
screen "01 Part Select" 480x800, template "Current Menu Selection"
   Button "B7" at 6,164 size 233x154; TextOff 'Text'
      on Press: function_b14e0dd5("pbs", 7)
      Visibility <- "[7]"
   Button "B6" at 6,323 size 233x154; TextOff 'Text'
      on Press: function_b14e0dd5("pbs", 6)
      Visibility <- "[6]"
   Button "B5" at 6,482 size 233x154; TextOff 'Text'
      on Press: function_b14e0dd5("pbs", 5)
      Visibility <- "[5]"
   Button "B4" at 6,641 size 233x154; TextOff 'Text'
      on Press: function_b14e0dd5("pbs", 4)
      Visibility <- "[4]"
   Button "B3" at 244,164 size 232x154; TextOff 'Text'
      on Press: function_b14e0dd5("pbs", 3)
      Visibility <- "[3]"
   Button "B2" at 244,323 size 232x154; TextOff 'Text'
      on Press: function_b14e0dd5("pbs", 2)
      Visibility <- "[2]"
   Button "B1" at 244,482 size 232x154; TextOff 'Text'
      on Press: function_b14e0dd5("pbs", 1)
      Visibility <- "[1]"
   Button "B0" at 244,641 size 232x154; TextOff 'Text'
      on Press: function_b14e0dd5("pbs", 0)
   IOField "B7 Label" at 6,164 size 233x154; FormatPattern ????????????????????????????????????????
      Appearance <- "[7]"
      ProcessValue <- "[7]"
      Visibility <- "[7]"
   IOField "B6 Label" at 6,323 size 233x154; FormatPattern ????????????????????????????????????????
      Appearance <- "[6]"
      ProcessValue <- "[6]"
      Visibility <- "[6]"
   IOField "B5 Label" at 6,482 size 233x154; FormatPattern ????????????????????????????????????????
      Appearance <- "[5]"
      ProcessValue <- "[5]"
      Visibility <- "[5]"
   IOField "B4 Label" at 6,641 size 233x154; FormatPattern ????????????????????????????????????????
      Appearance <- "[4]"
      ProcessValue <- "[4]"
      Visibility <- "[4]"
   IOField "B3 Label" at 244,164 size 232x154; FormatPattern ????????????????????????????????????????
      Appearance <- "[3]"
      ProcessValue <- "[3]"
      Visibility <- "[3]"
   IOField "B2 Label" at 244,323 size 232x154; FormatPattern ????????????????????????????????????????
      Appearance <- "[2]"
      ProcessValue <- "[2]"
      Visibility <- "[2]"
   IOField "B1 Label" at 244,482 size 232x154; FormatPattern ????????????????????????????????????????
      Appearance <- "[1]"
      ProcessValue <- "[1]"
      Visibility <- "[1]"
   IOField "B0 Label" at 244,641 size 232x154; FormatPattern ????????????????????????????????????????
      Appearance <- "[0]"
      ProcessValue <- "[0]"
      Visibility <- "[0]"

screen "02 Menu Select" 480x800, template "Current Menu Selection"
   Button "Top" at 375,164 size 100x101; TextOff 'Text'; PictureOff "basic panel top"
      on Press: function_b14e0dd5("pbs", 0)
      Appearance <- "[0]"
      Visibility <- "[0]"
   Button "Page Up" at 375,270 size 100x101; TextOff 'Text'; PictureOff "basic panel page up"
      on Press: function_b14e0dd5("pbs", 1)
      Visibility <- "[1]"
      Appearance <- "[1]"
   Button "Line Up" at 375,376 size 100x101; TextOff 'Text'; PictureOff "basic panel line up"
      on Press: function_b14e0dd5("pbs", 2)
      Appearance <- "[2]"
      Visibility <- "[2]"
   Button "Line Down" at 375,482 size 100x101; TextOff 'Text'; PictureOff "basic panel line down"
      on Press: function_b14e0dd5("pbs", 3)
      Visibility <- "[3]"
      Appearance <- "[3]"
   Button "Page Down" at 375,588 size 100x101; TextOff 'Text'; PictureOff "basic panel page down"
      on Press: function_b14e0dd5("pbs", 4)
      Appearance <- "[4]"
      Visibility <- "[4]"
   Button "Bottom" at 375,694 size 100x101; TextOff 'Text'; PictureOff "basic panel bottom"
      on Press: function_b14e0dd5("pbs", 5)
      Visibility <- "[5]"
      Appearance <- "[5]"
   IOField "brdrShortR00" at 5,164 size 365x101; FormatPattern 1
      Visibility <- "[6]"
      Appearance <- "[6]"
   IOField "brdrShortR01" at 5,270 size 365x101; FormatPattern 1
      Visibility <- "[7]"
      Appearance <- "[7]"
   IOField "brdrShortR02" at 5,376 size 365x101; FormatPattern 1
      Visibility <- "[8]"
      Appearance <- "[8]"
   IOField "brdrShortR03" at 5,482 size 365x101; FormatPattern 1
      Visibility <- "[9]"
      Appearance <- "[9]"
   IOField "brdrShortR04" at 5,588 size 365x101; FormatPattern 1
      Visibility <- "[10]"
      Appearance <- "[10]"
   IOField "brdrShortR05" at 5,694 size 365x101; FormatPattern 1
      Visibility <- "[11]"
      Appearance <- "[11]"
   Button "pbShortSelectR00" at 5,164 size 365x101; TextOff 'Text'
      on Release: ActivateScreen("01 Part Select", 0)
      on Press: function_b14e0dd5("pbs", 6)
   Button "pbShortSelectR01" at 5,270 size 365x101; TextOff 'Text'
      on Release: ActivateScreen("01 Part Select", 0)
      on Press: function_b14e0dd5("pbs", 7)
   Button "pbShortSelectR02" at 5,376 size 365x101; TextOff 'Text'
      on Release: ActivateScreen("01 Part Select", 0)
      on Press: function_b14e0dd5("pbs", 8)
   Button "pbShortSelectR03" at 5,482 size 365x101; TextOff 'Text'
      on Release: ActivateScreen("01 Part Select", 0)
      on Press: function_b14e0dd5("pbs", 9)
   Button "pbShortSelectR04" at 5,588 size 365x101; TextOff 'Text'
      on Release: ActivateScreen("01 Part Select", 0)
      on Press: function_b14e0dd5("pbs", 10)
   Button "pbShortSelectR05" at 5,694 size 365x101; TextOff 'Text'
      on Release: ActivateScreen("01 Part Select", 0)
      on Press: function_b14e0dd5("pbs", 11)
   IOField "brdrLongR00" at 5,164 size 470x101; FormatPattern 1
      Visibility <- "[18]"
   IOField "brdrLongR01" at 5,270 size 470x101; FormatPattern 1
      Visibility <- "[19]"
   IOField "brdrLongR02" at 5,376 size 470x101; FormatPattern 1
      Visibility <- "[20]"
   IOField "brdrLongR03" at 5,482 size 470x101; FormatPattern 1
      Visibility <- "[21]"
   IOField "brdrLongR04" at 5,588 size 470x101; FormatPattern 1
      Visibility <- "[22]"
   IOField "brdrLongR05" at 5,694 size 470x101; FormatPattern 1
      Visibility <- "[23]"
   Button "pbLongtSelectR00" at 5,164 size 470x101; TextOff 'Text'
      on Release: ActivateScreen("01 Part Select", 0)
      on Press: function_b14e0dd5("pbs", 6)
      Visibility <- "[18]"
   Button "pbLongtSelectR01" at 5,270 size 470x101; TextOff 'Text'
      on Release: ActivateScreen("01 Part Select", 0)
      on Press: function_b14e0dd5("pbs", 7)
      Visibility <- "[19]"
   Button "pbLongtSelectR02" at 5,376 size 470x101; TextOff 'Text'
      on Release: ActivateScreen("01 Part Select", 0)
      on Press: function_b14e0dd5("pbs", 8)
      Visibility <- "[20]"
   Button "pbLongtSelectR03" at 5,482 size 470x101; TextOff 'Text'
      on Release: ActivateScreen("01 Part Select", 0)
      on Press: function_b14e0dd5("pbs", 9)
      Visibility <- "[21]"
   Button "pbLongtSelectR04" at 5,588 size 470x101; TextOff 'Text'
      on Release: ActivateScreen("01 Part Select", 0)
      on Press: function_b14e0dd5("pbs", 10)
      Visibility <- "[22]"
   Button "pbLongtSelectR05" at 5,694 size 470x101; TextOff 'Text'
      on Release: ActivateScreen("01 Part Select", 0)
      on Press: function_b14e0dd5("pbs", 11)
      Visibility <- "[23]"
   IOField "iofLongtMenuSelectR00" at 42,166 size 430x97; FormatPattern ????????????????????????????????????????????????????????????
      Visibility <- "[18]"
      ProcessValue <- "[7]"
      Appearance <- "[18]"
   IOField "iofLongtMenuSelectR01" at 42,272 size 430x97; FormatPattern ????????????????????????????????????????????????????????????
      Visibility <- "[19]"
      ProcessValue <- "[9]"
      Appearance <- "[19]"
   IOField "iofLongtMenuSelectR02" at 42,378 size 430x97; FormatPattern ????????????????????????????????????????????????????????????
      Visibility <- "[20]"
      ProcessValue <- "[11]"
      Appearance <- "[20]"
   IOField "iofLongtMenuSelectR03" at 42,484 size 430x97; FormatPattern ????????????????????????????????????????????????????????????
      Visibility <- "[21]"
      ProcessValue <- "[13]"
      Appearance <- "[21]"
   IOField "iofLongtMenuSelectR04" at 42,590 size 430x97; FormatPattern ????????????????????????????????????????????????????????????
      Visibility <- "[22]"
      ProcessValue <- "[15]"
      Appearance <- "[22]"
   IOField "iofLongtMenuSelectR05" at 42,696 size 430x97; FormatPattern ????????????????????????????????????????????????????????????
      Visibility <- "[23]"
      ProcessValue <- "[17]"
      Appearance <- "[22]"
   IOField "iofLongLabelR00" at 7,166 size 35x97; FormatPattern ????????????????????????????????????????
      Visibility <- "[18]"
      ProcessValue <- "[6]"
      Appearance <- "[18]"
   IOField "iofLongLabelR01" at 7,272 size 35x97; FormatPattern ????????????????????????????????????????
      Appearance <- "[19]"
      ProcessValue <- "[8]"
      Visibility <- "[19]"
   IOField "iofLongLabelR02" at 7,378 size 35x97; FormatPattern ????????????????????????????????????????
      Appearance <- "[20]"
      ProcessValue <- "[10]"
      Visibility <- "[20]"
   IOField "iofLongLabelR03" at 7,484 size 35x97; FormatPattern ????????????????????????????????????????
      Appearance <- "[21]"
      ProcessValue <- "[12]"
      Visibility <- "[21]"
   IOField "iofLongLabelR04" at 7,590 size 35x97; FormatPattern ????????????????????????????????????????
      Visibility <- "[22]"
      ProcessValue <- "[14]"
      Appearance <- "[22]"
   IOField "iofLongtLabelR05" at 7,696 size 35x97; FormatPattern ????????????????????????????????????????
      Appearance <- "[23]"
      ProcessValue <- "[16]"
      Visibility <- "[23]"
   IOField "iofShortMenuSelectR00" at 42,166 size 325x97; FormatPattern ????????????????????????????????????????????????????????????
      Visibility <- "[6]"
      ProcessValue <- "[7]"
      Appearance <- "[6]"
   IOField "iofShortMenuSelectR01" at 42,272 size 325x97; FormatPattern ????????????????????????????????????????????????????????????
      Visibility <- "[7]"
      ProcessValue <- "[9]"
      Appearance <- "[7]"
   IOField "iofShortMenuSelectR02" at 42,378 size 325x97; FormatPattern ????????????????????????????????????????????????????????????
      Visibility <- "[8]"
      ProcessValue <- "[11]"
      Appearance <- "[8]"
   IOField "iofShortMenuSelectR03" at 42,484 size 325x97; FormatPattern ????????????????????????????????????????????????????????????
      Visibility <- "[9]"
      ProcessValue <- "[13]"
      Appearance <- "[9]"
   IOField "iofShortMenuSelectR04" at 42,590 size 325x97; FormatPattern ????????????????????????????????????????????????????????????
      Visibility <- "[10]"
      ProcessValue <- "[15]"
      Appearance <- "[10]"
   IOField "iofShortMenuSelectR05" at 42,696 size 325x97; FormatPattern ????????????????????????????????????????????????????????????
      Visibility <- "[11]"
      ProcessValue <- "[17]"
      Appearance <- "[11]"
   IOField "iofShortLabelR00" at 7,166 size 35x97; FormatPattern ????????????????????????????????????????
      Appearance <- "[6]"
      ProcessValue <- "[6]"
      Visibility <- "[6]"
   IOField "iofShortLabelR01" at 7,272 size 35x97; FormatPattern ????????????????????????????????????????
      Appearance <- "[7]"
      ProcessValue <- "[8]"
      Visibility <- "[7]"
   IOField "iofShortLabelR02" at 7,378 size 35x97; FormatPattern ????????????????????????????????????????
      Appearance <- "[8]"
      ProcessValue <- "[10]"
      Visibility <- "[8]"
   IOField "iofShortLabelR03" at 7,484 size 35x97; FormatPattern ????????????????????????????????????????
      Appearance <- "[9]"
      ProcessValue <- "[12]"
      Visibility <- "[9]"
   IOField "iofShortLabelR04" at 7,590 size 35x97; FormatPattern ????????????????????????????????????????
      Appearance <- "[10]"
      ProcessValue <- "[14]"
      Visibility <- "[10]"
   IOField "iofShorttLabelR05" at 7,696 size 35x97; FormatPattern ????????????????????????????????????????
      Appearance <- "[11]"
      ProcessValue <- "[16]"
      Visibility <- "[11]"

Template "Current Menu Selection" 480x800
   IOField "Menu Select Label" at 6,5 size 470x154; FormatPattern ????????????????????????????????????????????????????????????
      Appearance <- "[0]"
      Visibility <- "[0]"
      ProcessValue <- "[0]"
   Button "PB Menu Select" at 6,5 size 470x154; TextOff 'Text'
      on Release: ActivateScreen("02 Menu Select", 0)
      on Press: function_b14e0dd5("pb", 0)
*)

(* ===== HMI "HMI_RT_6" =====
system functions are stored by id; their names below are inferred from use
connection "cv01": ETHERNET, SMART_S7_1500_OMS

HMI tags "Default tag table"
   "station" : HMIS: Compressed = PLC "HMI Stations".me[0] AT %DB1.DBW0, 100 ms

screen "01 Part Select" 480x800, template "Current Menu Selection"
   Button "B7" at 6,164 size 233x154; TextOff 'Text'
      on Press: function_b14e0dd5("pbs", 7)
      Visibility <- "[7]"
   Button "B6" at 6,323 size 233x154; TextOff 'Text'
      on Press: function_b14e0dd5("pbs", 6)
      Visibility <- "[6]"
   Button "B5" at 6,482 size 233x154; TextOff 'Text'
      on Press: function_b14e0dd5("pbs", 5)
      Visibility <- "[5]"
   Button "B4" at 6,641 size 233x154; TextOff 'Text'
      on Press: function_b14e0dd5("pbs", 4)
      Visibility <- "[4]"
   Button "B3" at 244,164 size 232x154; TextOff 'Text'
      on Press: function_b14e0dd5("pbs", 3)
      Visibility <- "[3]"
   Button "B2" at 244,323 size 232x154; TextOff 'Text'
      on Press: function_b14e0dd5("pbs", 2)
      Visibility <- "[2]"
   Button "B1" at 244,482 size 232x154; TextOff 'Text'
      on Press: function_b14e0dd5("pbs", 1)
      Visibility <- "[1]"
   Button "B0" at 244,641 size 232x154; TextOff 'Text'
      on Press: function_b14e0dd5("pbs", 0)
   IOField "B7 Label" at 6,164 size 233x154; FormatPattern ????????????????????????????????????????
      Appearance <- "[7]"
      ProcessValue <- "[7]"
      Visibility <- "[7]"
   IOField "B6 Label" at 6,323 size 233x154; FormatPattern ????????????????????????????????????????
      Appearance <- "[6]"
      ProcessValue <- "[6]"
      Visibility <- "[6]"
   IOField "B5 Label" at 6,482 size 233x154; FormatPattern ????????????????????????????????????????
      Appearance <- "[5]"
      ProcessValue <- "[5]"
      Visibility <- "[5]"
   IOField "B4 Label" at 6,641 size 233x154; FormatPattern ????????????????????????????????????????
      Appearance <- "[4]"
      ProcessValue <- "[4]"
      Visibility <- "[4]"
   IOField "B3 Label" at 244,164 size 232x154; FormatPattern ????????????????????????????????????????
      Appearance <- "[3]"
      ProcessValue <- "[3]"
      Visibility <- "[3]"
   IOField "B2 Label" at 244,323 size 232x154; FormatPattern ????????????????????????????????????????
      Appearance <- "[2]"
      ProcessValue <- "[2]"
      Visibility <- "[2]"
   IOField "B1 Label" at 244,482 size 232x154; FormatPattern ????????????????????????????????????????
      Appearance <- "[1]"
      ProcessValue <- "[1]"
      Visibility <- "[1]"
   IOField "B0 Label" at 244,641 size 232x154; FormatPattern ????????????????????????????????????????
      Appearance <- "[0]"
      ProcessValue <- "[0]"
      Visibility <- "[0]"
   TextField "B7 BG" at 6,164 size 233x154; Text '1'

screen "02 Menu Select" 480x800, template "Current Menu Selection"
   Button "Top" at 375,164 size 100x101; TextOff 'Text'; PictureOff "basic panel top"
      on Press: function_b14e0dd5("pbs", 0)
      Appearance <- "[0]"
      Visibility <- "[0]"
   Button "Page Up" at 375,270 size 100x101; TextOff 'Text'; PictureOff "basic panel page up"
      on Press: function_b14e0dd5("pbs", 1)
      Visibility <- "[1]"
      Appearance <- "[1]"
   Button "Line Up" at 375,376 size 100x101; TextOff 'Text'; PictureOff "basic panel line up"
      on Press: function_b14e0dd5("pbs", 2)
      Appearance <- "[2]"
      Visibility <- "[2]"
   Button "Line Down" at 375,482 size 100x101; TextOff 'Text'; PictureOff "basic panel line down"
      on Press: function_b14e0dd5("pbs", 3)
      Visibility <- "[3]"
      Appearance <- "[3]"
   Button "Page Down" at 375,588 size 100x101; TextOff 'Text'; PictureOff "basic panel page down"
      on Press: function_b14e0dd5("pbs", 4)
      Appearance <- "[4]"
      Visibility <- "[4]"
   Button "Bottom" at 375,694 size 100x101; TextOff 'Text'; PictureOff "basic panel bottom"
      on Press: function_b14e0dd5("pbs", 5)
      Visibility <- "[5]"
      Appearance <- "[5]"
   IOField "brdrShortR00" at 5,164 size 365x101; FormatPattern 1
      Visibility <- "[6]"
      Appearance <- "[6]"
   IOField "brdrShortR01" at 5,270 size 365x101; FormatPattern 1
      Visibility <- "[7]"
      Appearance <- "[7]"
   IOField "brdrShortR02" at 5,376 size 365x101; FormatPattern 1
      Visibility <- "[8]"
      Appearance <- "[8]"
   IOField "brdrShortR03" at 5,482 size 365x101; FormatPattern 1
      Visibility <- "[9]"
      Appearance <- "[9]"
   IOField "brdrShortR04" at 5,588 size 365x101; FormatPattern 1
      Visibility <- "[10]"
      Appearance <- "[10]"
   IOField "brdrShortR05" at 5,694 size 365x101; FormatPattern 1
      Visibility <- "[11]"
      Appearance <- "[11]"
   Button "pbShortSelectR00" at 5,164 size 365x101; TextOff 'Text'
      on Release: ActivateScreen("01 Part Select", 0)
      on Press: function_b14e0dd5("pbs", 6)
   Button "pbShortSelectR01" at 5,270 size 365x101; TextOff 'Text'
      on Release: ActivateScreen("01 Part Select", 0)
      on Press: function_b14e0dd5("pbs", 7)
   Button "pbShortSelectR02" at 5,376 size 365x101; TextOff 'Text'
      on Release: ActivateScreen("01 Part Select", 0)
      on Press: function_b14e0dd5("pbs", 8)
   Button "pbShortSelectR03" at 5,482 size 365x101; TextOff 'Text'
      on Release: ActivateScreen("01 Part Select", 0)
      on Press: function_b14e0dd5("pbs", 9)
   Button "pbShortSelectR04" at 5,588 size 365x101; TextOff 'Text'
      on Release: ActivateScreen("01 Part Select", 0)
      on Press: function_b14e0dd5("pbs", 10)
   Button "pbShortSelectR05" at 5,694 size 365x101; TextOff 'Text'
      on Release: ActivateScreen("01 Part Select", 0)
      on Press: function_b14e0dd5("pbs", 11)
   IOField "brdrLongR00" at 5,164 size 470x101; FormatPattern 1
      Visibility <- "[18]"
   IOField "brdrLongR01" at 5,270 size 470x101; FormatPattern 1
      Visibility <- "[19]"
   IOField "brdrLongR02" at 5,376 size 470x101; FormatPattern 1
      Visibility <- "[20]"
   IOField "brdrLongR03" at 5,482 size 470x101; FormatPattern 1
      Visibility <- "[21]"
   IOField "brdrLongR04" at 5,588 size 470x101; FormatPattern 1
      Visibility <- "[22]"
   IOField "brdrLongR05" at 5,694 size 470x101; FormatPattern 1
      Visibility <- "[23]"
   Button "pbLongtSelectR00" at 5,164 size 470x101; TextOff 'Text'
      on Release: ActivateScreen("01 Part Select", 0)
      on Press: function_b14e0dd5("pbs", 6)
      Visibility <- "[18]"
   Button "pbLongtSelectR01" at 5,270 size 470x101; TextOff 'Text'
      on Release: ActivateScreen("01 Part Select", 0)
      on Press: function_b14e0dd5("pbs", 7)
      Visibility <- "[19]"
   Button "pbLongtSelectR02" at 5,376 size 470x101; TextOff 'Text'
      on Release: ActivateScreen("01 Part Select", 0)
      on Press: function_b14e0dd5("pbs", 8)
      Visibility <- "[20]"
   Button "pbLongtSelectR03" at 5,482 size 470x101; TextOff 'Text'
      on Release: ActivateScreen("01 Part Select", 0)
      on Press: function_b14e0dd5("pbs", 9)
      Visibility <- "[21]"
   Button "pbLongtSelectR04" at 5,588 size 470x101; TextOff 'Text'
      on Release: ActivateScreen("01 Part Select", 0)
      on Press: function_b14e0dd5("pbs", 10)
      Visibility <- "[22]"
   Button "pbLongtSelectR05" at 5,694 size 470x101; TextOff 'Text'
      on Release: ActivateScreen("01 Part Select", 0)
      on Press: function_b14e0dd5("pbs", 11)
      Visibility <- "[23]"
   IOField "iofLongtMenuSelectR00" at 42,166 size 430x97; FormatPattern ????????????????????????????????????????????????????????????
      Visibility <- "[18]"
      ProcessValue <- "[7]"
      Appearance <- "[18]"
   IOField "iofLongtMenuSelectR01" at 42,272 size 430x97; FormatPattern ????????????????????????????????????????????????????????????
      Visibility <- "[19]"
      ProcessValue <- "[9]"
      Appearance <- "[19]"
   IOField "iofLongtMenuSelectR02" at 42,378 size 430x97; FormatPattern ????????????????????????????????????????????????????????????
      Visibility <- "[20]"
      ProcessValue <- "[11]"
      Appearance <- "[20]"
   IOField "iofLongtMenuSelectR03" at 42,484 size 430x97; FormatPattern ????????????????????????????????????????????????????????????
      Visibility <- "[21]"
      ProcessValue <- "[13]"
      Appearance <- "[21]"
   IOField "iofLongtMenuSelectR04" at 42,590 size 430x97; FormatPattern ????????????????????????????????????????????????????????????
      Visibility <- "[22]"
      ProcessValue <- "[15]"
      Appearance <- "[22]"
   IOField "iofLongtMenuSelectR05" at 42,696 size 430x97; FormatPattern ????????????????????????????????????????????????????????????
      Visibility <- "[23]"
      ProcessValue <- "[17]"
      Appearance <- "[22]"
   IOField "iofLongLabelR00" at 7,166 size 35x97; FormatPattern ????????????????????????????????????????
      Visibility <- "[18]"
      ProcessValue <- "[6]"
      Appearance <- "[18]"
   IOField "iofLongLabelR01" at 7,272 size 35x97; FormatPattern ????????????????????????????????????????
      Appearance <- "[19]"
      ProcessValue <- "[8]"
      Visibility <- "[19]"
   IOField "iofLongLabelR02" at 7,378 size 35x97; FormatPattern ????????????????????????????????????????
      Appearance <- "[20]"
      ProcessValue <- "[10]"
      Visibility <- "[20]"
   IOField "iofLongLabelR03" at 7,484 size 35x97; FormatPattern ????????????????????????????????????????
      Appearance <- "[21]"
      ProcessValue <- "[12]"
      Visibility <- "[21]"
   IOField "iofLongLabelR04" at 7,590 size 35x97; FormatPattern ????????????????????????????????????????
      Visibility <- "[22]"
      ProcessValue <- "[14]"
      Appearance <- "[22]"
   IOField "iofLongtLabelR05" at 7,696 size 35x97; FormatPattern ????????????????????????????????????????
      Appearance <- "[23]"
      ProcessValue <- "[16]"
      Visibility <- "[23]"
   IOField "iofShortMenuSelectR00" at 42,166 size 325x97; FormatPattern ????????????????????????????????????????????????????????????
      Visibility <- "[6]"
      ProcessValue <- "[7]"
      Appearance <- "[6]"
   IOField "iofShortMenuSelectR01" at 42,272 size 325x97; FormatPattern ????????????????????????????????????????????????????????????
      Visibility <- "[7]"
      ProcessValue <- "[9]"
      Appearance <- "[7]"
   IOField "iofShortMenuSelectR02" at 42,378 size 325x97; FormatPattern ????????????????????????????????????????????????????????????
      Visibility <- "[8]"
      ProcessValue <- "[11]"
      Appearance <- "[8]"
   IOField "iofShortMenuSelectR03" at 42,484 size 325x97; FormatPattern ????????????????????????????????????????????????????????????
      Visibility <- "[9]"
      ProcessValue <- "[13]"
      Appearance <- "[9]"
   IOField "iofShortMenuSelectR04" at 42,590 size 325x97; FormatPattern ????????????????????????????????????????????????????????????
      Visibility <- "[10]"
      ProcessValue <- "[15]"
      Appearance <- "[10]"
   IOField "iofShortMenuSelectR05" at 42,696 size 325x97; FormatPattern ????????????????????????????????????????????????????????????
      Visibility <- "[11]"
      ProcessValue <- "[17]"
      Appearance <- "[11]"
   IOField "iofShortLabelR00" at 7,166 size 35x97; FormatPattern ????????????????????????????????????????
      Appearance <- "[6]"
      ProcessValue <- "[6]"
      Visibility <- "[6]"
   IOField "iofShortLabelR01" at 7,272 size 35x97; FormatPattern ????????????????????????????????????????
      Appearance <- "[7]"
      ProcessValue <- "[8]"
      Visibility <- "[7]"
   IOField "iofShortLabelR02" at 7,378 size 35x97; FormatPattern ????????????????????????????????????????
      Appearance <- "[8]"
      ProcessValue <- "[10]"
      Visibility <- "[8]"
   IOField "iofShortLabelR03" at 7,484 size 35x97; FormatPattern ????????????????????????????????????????
      Appearance <- "[9]"
      ProcessValue <- "[12]"
      Visibility <- "[9]"
   IOField "iofShortLabelR04" at 7,590 size 35x97; FormatPattern ????????????????????????????????????????
      Appearance <- "[10]"
      ProcessValue <- "[14]"
      Visibility <- "[10]"
   IOField "iofShorttLabelR05" at 7,696 size 35x97; FormatPattern ????????????????????????????????????????
      Appearance <- "[11]"
      ProcessValue <- "[16]"
      Visibility <- "[11]"

Template "Current Menu Selection" 480x800
   IOField "Menu Select Label" at 6,5 size 470x154; FormatPattern ????????????????????????????????????????????????????????????
      Appearance <- "[0]"
      Visibility <- "[0]"
      ProcessValue <- "[0]"
   Button "PB Menu Select" at 6,5 size 470x154; TextOff 'Text'
      on Release: ActivateScreen("02 Menu Select", 0)
      on Press: function_b14e0dd5("pb", 0)
*)

(* ===== HMI "HMI_RT_7" =====
system functions are stored by id; their names below are inferred from use
connection "pc01": ETHERNET, SMART_S7_1500_OMS

HMI tags "Default tag table"
   "station" : HMIS: Compressed = PLC "HMI Stations".me[4] AT %DB1.DBW0, 100 ms

screen "01 Part Select" 480x800, template "Current Menu Selection"
   Button "B7" at 6,164 size 233x154; TextOff 'Text'
      on Press: function_b14e0dd5("pbs", 7)
      Visibility <- "[7]"
   Button "B6" at 6,323 size 233x154; TextOff 'Text'
      on Press: function_b14e0dd5("pbs", 6)
      Visibility <- "[6]"
   Button "B5" at 6,482 size 233x154; TextOff 'Text'
      on Press: function_b14e0dd5("pbs", 5)
      Visibility <- "[5]"
   Button "B4" at 6,641 size 233x154; TextOff 'Text'
      on Press: function_b14e0dd5("pbs", 4)
      Visibility <- "[4]"
   Button "B3" at 244,164 size 232x154; TextOff 'Text'
      on Press: function_b14e0dd5("pbs", 3)
      Visibility <- "[3]"
   Button "B2" at 244,323 size 232x154; TextOff 'Text'
      on Press: function_b14e0dd5("pbs", 2)
      Visibility <- "[2]"
   Button "B1" at 244,482 size 232x154; TextOff 'Text'
      on Press: function_b14e0dd5("pbs", 1)
      Visibility <- "[1]"
   Button "B0" at 244,641 size 232x154; TextOff 'Text'
      on Press: function_b14e0dd5("pbs", 0)
   IOField "B7 Label" at 6,164 size 233x154; FormatPattern ????????????????????????????????????????
      Appearance <- "[7]"
      ProcessValue <- "[7]"
      Visibility <- "[7]"
   IOField "B6 Label" at 6,323 size 233x154; FormatPattern ????????????????????????????????????????
      Appearance <- "[6]"
      ProcessValue <- "[6]"
      Visibility <- "[6]"
   IOField "B5 Label" at 6,482 size 233x154; FormatPattern ????????????????????????????????????????
      Appearance <- "[5]"
      ProcessValue <- "[5]"
      Visibility <- "[5]"
   IOField "B4 Label" at 6,641 size 233x154; FormatPattern ????????????????????????????????????????
      Appearance <- "[4]"
      ProcessValue <- "[4]"
      Visibility <- "[4]"
   IOField "B3 Label" at 244,164 size 232x154; FormatPattern ????????????????????????????????????????
      Appearance <- "[3]"
      ProcessValue <- "[3]"
      Visibility <- "[3]"
   IOField "B2 Label" at 244,323 size 232x154; FormatPattern ????????????????????????????????????????
      Appearance <- "[2]"
      ProcessValue <- "[2]"
      Visibility <- "[2]"
   IOField "B1 Label" at 244,482 size 232x154; FormatPattern ????????????????????????????????????????
      Appearance <- "[1]"
      ProcessValue <- "[1]"
      Visibility <- "[1]"
   IOField "B0 Label" at 244,641 size 232x154; FormatPattern ????????????????????????????????????????
      Appearance <- "[0]"
      ProcessValue <- "[0]"
      Visibility <- "[0]"

screen "02 Menu Select" 480x800, template "Current Menu Selection"
   Button "Top" at 375,164 size 100x101; TextOff 'Text'; PictureOff "basic panel top"
      on Press: function_b14e0dd5("pbs", 0)
      Appearance <- "[0]"
      Visibility <- "[0]"
   Button "Page Up" at 375,270 size 100x101; TextOff 'Text'; PictureOff "basic panel page up"
      on Press: function_b14e0dd5("pbs", 1)
      Visibility <- "[1]"
      Appearance <- "[1]"
   Button "Line Up" at 375,376 size 100x101; TextOff 'Text'; PictureOff "basic panel line up"
      on Press: function_b14e0dd5("pbs", 2)
      Appearance <- "[2]"
      Visibility <- "[2]"
   Button "Line Down" at 375,482 size 100x101; TextOff 'Text'; PictureOff "basic panel line down"
      on Press: function_b14e0dd5("pbs", 3)
      Visibility <- "[3]"
      Appearance <- "[3]"
   Button "Page Down" at 375,588 size 100x101; TextOff 'Text'; PictureOff "basic panel page down"
      on Press: function_b14e0dd5("pbs", 4)
      Appearance <- "[4]"
      Visibility <- "[4]"
   Button "Bottom" at 375,694 size 100x101; TextOff 'Text'; PictureOff "basic panel bottom"
      on Press: function_b14e0dd5("pbs", 5)
      Visibility <- "[5]"
      Appearance <- "[5]"
   IOField "brdrShortR00" at 5,164 size 365x101; FormatPattern 1
      Visibility <- "[6]"
      Appearance <- "[6]"
   IOField "brdrShortR01" at 5,270 size 365x101; FormatPattern 1
      Visibility <- "[7]"
      Appearance <- "[7]"
   IOField "brdrShortR02" at 5,376 size 365x101; FormatPattern 1
      Visibility <- "[8]"
      Appearance <- "[8]"
   IOField "brdrShortR03" at 5,482 size 365x101; FormatPattern 1
      Visibility <- "[9]"
      Appearance <- "[9]"
   IOField "brdrShortR04" at 5,588 size 365x101; FormatPattern 1
      Visibility <- "[10]"
      Appearance <- "[10]"
   IOField "brdrShortR05" at 5,694 size 365x101; FormatPattern 1
      Visibility <- "[11]"
      Appearance <- "[11]"
   Button "pbShortSelectR00" at 5,164 size 365x101; TextOff 'Text'
      on Release: ActivateScreen("01 Part Select", 0)
      on Press: function_b14e0dd5("pbs", 6)
   Button "pbShortSelectR01" at 5,270 size 365x101; TextOff 'Text'
      on Release: ActivateScreen("01 Part Select", 0)
      on Press: function_b14e0dd5("pbs", 7)
   Button "pbShortSelectR02" at 5,376 size 365x101; TextOff 'Text'
      on Release: ActivateScreen("01 Part Select", 0)
      on Press: function_b14e0dd5("pbs", 8)
   Button "pbShortSelectR03" at 5,482 size 365x101; TextOff 'Text'
      on Release: ActivateScreen("01 Part Select", 0)
      on Press: function_b14e0dd5("pbs", 9)
   Button "pbShortSelectR04" at 5,588 size 365x101; TextOff 'Text'
      on Release: ActivateScreen("01 Part Select", 0)
      on Press: function_b14e0dd5("pbs", 10)
   Button "pbShortSelectR05" at 5,694 size 365x101; TextOff 'Text'
      on Release: ActivateScreen("01 Part Select", 0)
      on Press: function_b14e0dd5("pbs", 11)
   IOField "brdrLongR00" at 5,164 size 470x101; FormatPattern 1
      Visibility <- "[18]"
   IOField "brdrLongR01" at 5,270 size 470x101; FormatPattern 1
      Visibility <- "[19]"
   IOField "brdrLongR02" at 5,376 size 470x101; FormatPattern 1
      Visibility <- "[20]"
   IOField "brdrLongR03" at 5,482 size 470x101; FormatPattern 1
      Visibility <- "[21]"
   IOField "brdrLongR04" at 5,588 size 470x101; FormatPattern 1
      Visibility <- "[22]"
   IOField "brdrLongR05" at 5,694 size 470x101; FormatPattern 1
      Visibility <- "[23]"
   Button "pbLongtSelectR00" at 5,164 size 470x101; TextOff 'Text'
      on Release: ActivateScreen("01 Part Select", 0)
      on Press: function_b14e0dd5("pbs", 6)
      Visibility <- "[18]"
   Button "pbLongtSelectR01" at 5,270 size 470x101; TextOff 'Text'
      on Release: ActivateScreen("01 Part Select", 0)
      on Press: function_b14e0dd5("pbs", 7)
      Visibility <- "[19]"
   Button "pbLongtSelectR02" at 5,376 size 470x101; TextOff 'Text'
      on Release: ActivateScreen("01 Part Select", 0)
      on Press: function_b14e0dd5("pbs", 8)
      Visibility <- "[20]"
   Button "pbLongtSelectR03" at 5,482 size 470x101; TextOff 'Text'
      on Release: ActivateScreen("01 Part Select", 0)
      on Press: function_b14e0dd5("pbs", 9)
      Visibility <- "[21]"
   Button "pbLongtSelectR04" at 5,588 size 470x101; TextOff 'Text'
      on Release: ActivateScreen("01 Part Select", 0)
      on Press: function_b14e0dd5("pbs", 10)
      Visibility <- "[22]"
   Button "pbLongtSelectR05" at 5,694 size 470x101; TextOff 'Text'
      on Release: ActivateScreen("01 Part Select", 0)
      on Press: function_b14e0dd5("pbs", 11)
      Visibility <- "[23]"
   IOField "iofLongtMenuSelectR00" at 42,166 size 430x97; FormatPattern ????????????????????????????????????????????????????????????
      Visibility <- "[18]"
      ProcessValue <- "[7]"
      Appearance <- "[18]"
   IOField "iofLongtMenuSelectR01" at 42,272 size 430x97; FormatPattern ????????????????????????????????????????????????????????????
      Visibility <- "[19]"
      ProcessValue <- "[9]"
      Appearance <- "[19]"
   IOField "iofLongtMenuSelectR02" at 42,378 size 430x97; FormatPattern ????????????????????????????????????????????????????????????
      Visibility <- "[20]"
      ProcessValue <- "[11]"
      Appearance <- "[20]"
   IOField "iofLongtMenuSelectR03" at 42,484 size 430x97; FormatPattern ????????????????????????????????????????????????????????????
      Visibility <- "[21]"
      ProcessValue <- "[13]"
      Appearance <- "[21]"
   IOField "iofLongtMenuSelectR04" at 42,590 size 430x97; FormatPattern ????????????????????????????????????????????????????????????
      Visibility <- "[22]"
      ProcessValue <- "[15]"
      Appearance <- "[22]"
   IOField "iofLongtMenuSelectR05" at 42,696 size 430x97; FormatPattern ????????????????????????????????????????????????????????????
      Visibility <- "[23]"
      ProcessValue <- "[17]"
      Appearance <- "[22]"
   IOField "iofLongLabelR00" at 7,166 size 35x97; FormatPattern ????????????????????????????????????????
      Visibility <- "[18]"
      ProcessValue <- "[6]"
      Appearance <- "[18]"
   IOField "iofLongLabelR01" at 7,272 size 35x97; FormatPattern ????????????????????????????????????????
      Appearance <- "[19]"
      ProcessValue <- "[8]"
      Visibility <- "[19]"
   IOField "iofLongLabelR02" at 7,378 size 35x97; FormatPattern ????????????????????????????????????????
      Appearance <- "[20]"
      ProcessValue <- "[10]"
      Visibility <- "[20]"
   IOField "iofLongLabelR03" at 7,484 size 35x97; FormatPattern ????????????????????????????????????????
      Appearance <- "[21]"
      ProcessValue <- "[12]"
      Visibility <- "[21]"
   IOField "iofLongLabelR04" at 7,590 size 35x97; FormatPattern ????????????????????????????????????????
      Visibility <- "[22]"
      ProcessValue <- "[14]"
      Appearance <- "[22]"
   IOField "iofLongtLabelR05" at 7,696 size 35x97; FormatPattern ????????????????????????????????????????
      Appearance <- "[23]"
      ProcessValue <- "[16]"
      Visibility <- "[23]"
   IOField "iofShortMenuSelectR00" at 42,166 size 325x97; FormatPattern ????????????????????????????????????????????????????????????
      Visibility <- "[6]"
      ProcessValue <- "[7]"
      Appearance <- "[6]"
   IOField "iofShortMenuSelectR01" at 42,272 size 325x97; FormatPattern ????????????????????????????????????????????????????????????
      Visibility <- "[7]"
      ProcessValue <- "[9]"
      Appearance <- "[7]"
   IOField "iofShortMenuSelectR02" at 42,378 size 325x97; FormatPattern ????????????????????????????????????????????????????????????
      Visibility <- "[8]"
      ProcessValue <- "[11]"
      Appearance <- "[8]"
   IOField "iofShortMenuSelectR03" at 42,484 size 325x97; FormatPattern ????????????????????????????????????????????????????????????
      Visibility <- "[9]"
      ProcessValue <- "[13]"
      Appearance <- "[9]"
   IOField "iofShortMenuSelectR04" at 42,590 size 325x97; FormatPattern ????????????????????????????????????????????????????????????
      Visibility <- "[10]"
      ProcessValue <- "[15]"
      Appearance <- "[10]"
   IOField "iofShortMenuSelectR05" at 42,696 size 325x97; FormatPattern ????????????????????????????????????????????????????????????
      Visibility <- "[11]"
      ProcessValue <- "[17]"
      Appearance <- "[11]"
   IOField "iofShortLabelR00" at 7,166 size 35x97; FormatPattern ????????????????????????????????????????
      Appearance <- "[6]"
      ProcessValue <- "[6]"
      Visibility <- "[6]"
   IOField "iofShortLabelR01" at 7,272 size 35x97; FormatPattern ????????????????????????????????????????
      Appearance <- "[7]"
      ProcessValue <- "[8]"
      Visibility <- "[7]"
   IOField "iofShortLabelR02" at 7,378 size 35x97; FormatPattern ????????????????????????????????????????
      Appearance <- "[8]"
      ProcessValue <- "[10]"
      Visibility <- "[8]"
   IOField "iofShortLabelR03" at 7,484 size 35x97; FormatPattern ????????????????????????????????????????
      Appearance <- "[9]"
      ProcessValue <- "[12]"
      Visibility <- "[9]"
   IOField "iofShortLabelR04" at 7,590 size 35x97; FormatPattern ????????????????????????????????????????
      Appearance <- "[10]"
      ProcessValue <- "[14]"
      Visibility <- "[10]"
   IOField "iofShorttLabelR05" at 7,696 size 35x97; FormatPattern ????????????????????????????????????????
      Appearance <- "[11]"
      ProcessValue <- "[16]"
      Visibility <- "[11]"

Template "Current Menu Selection" 480x800
   IOField "Menu Select Label" at 6,5 size 470x154; FormatPattern ????????????????????????????????????????????????????????????
      Appearance <- "[0]"
      Visibility <- "[0]"
      ProcessValue <- "[0]"
   Button "PB Menu Select" at 6,5 size 470x154; TextOff 'Text'
      on Release: ActivateScreen("02 Menu Select", 0)
      on Press: function_b14e0dd5("pb", 0)
*)